
screen "2005_ProNet temperature input" 1280x800, template "Navigation"
   Group "Group" at 118,204 size 1041x515
   TextField "Text field_3" at 172,348 size 56x25; Text 'Mode'
   TextField "Text field_4" at 172,388 size 56x25; Text 'Mode'
   TextField "Text field_5" at 172,430 size 105x25; Text 'Value_10V'
   TextField "Text field_6" at 172,470 size 139x25; Text 'Tank_Average'
   TextField "Text field_7" at 457,550 size 254x25; Text '0:0.. 5 V; 1: -5.. +5 V;'
   TextField "Text field_8" at 702,550 size 308x25; Text '2:0.. 10 V; 3: -10 V.. +10 V;'
   TextField "Text field_9" at 222,550 size 56x25; Text 'Mode'
   TextField "Text field_11" at 222,606 size 105x25; Text 'Value_10V'
   TextField "Text field_12" at 222,634 size 139x25; Text 'Tank_Average'
   TextField "Text field_14" at 457,606 size 366x25; Text 'Max Value for input 10V or 138.5 ohm'
   TextField "Text field_15" at 456,634 size 222x25; Text 'Time for average [ms]'
   TextField "Text field_16" at 373,302 size 46x25; Text '1'
   TextField "Text field_17" at 469,302 size 46x25; Text '2'
   TextField "Text field_18" at 565,302 size 46x25; Text '3'
   TextField "Text field_19" at 661,302 size 46x25; Text '4'
   TextField "Text field_20" at 757,302 size 46x25; Text '5'
   TextField "Text field_21" at 853,302 size 46x25; Text '6'
   TextField "Text field_22" at 949,302 size 46x25; Text '7'
   TextField "Text field_23" at 1045,302 size 46x25; Text '8'
   SymbolicIOField "Symbolic I/O field_5" at 326,104 size 451x32; TextOn '1'; TextOff '0'; TextList "Pronet_Analog_Input"
      ProcessValue <- "PN_AI_SetIndex"
   Button "b_Incress_PronetAnalogInput" at 787,104 size 46x32; TextOff 'Text'; PictureOff "NEXT"
      on Press: function_dd21b452("PN_AI_SetIndex", 1)
   Button "b_Decress_PronetAnalogInput" at 270,104 size 46x32; TextOff 'Text'; PictureOff "BEFORE"
      on Press: function_b9b71300("PN_AI_SetIndex", 1)
   Button "Button_1" at 1017,244 size 96x32; TextOff 'Active'
      on Press: InvertBit("PN_AI_Module{0}_AIResistive_8_Active")
      Appearance <- "PN_AI_Module{0}_AIResistive_8_Active"
   TextField "Text field_1" at 428,145 size 247x29; Text 'ProNet Configuration'
   IOField "Pronet_Analog_Input/Mode1" at 341,344 size 80x32; FormatPattern 9999999
      ProcessValue <- "PN_AI_Module{0}_AI8_X14_0_Data_Data[1]_Betriebsart"
   IOField "I/O field_2" at 437,344 size 80x32; FormatPattern 9999999
      ProcessValue <- "PN_AI_Module{0}_AI8_X14_0_Data_Data[2]_Betriebsart"
   IOField "I/O field_3" at 533,344 size 80x32; FormatPattern 9999999
      ProcessValue <- "PN_AI_Module{0}_AI8_X14_0_Data_Data[3]_Betriebsart"
   IOField "I/O field_4" at 629,344 size 80x32; FormatPattern 9999999
      ProcessValue <- "PN_AI_Module{0}_AI8_X14_0_Data_Data[4]_Betriebsart"
   IOField "I/O field_5" at 725,344 size 80x32; FormatPattern 9999999
      ProcessValue <- "PN_AI_Module{0}_AI8_X14_0_Data_Data[5]_Betriebsart"
   IOField "I/O field_6" at 821,344 size 80x32; FormatPattern 9999999
      ProcessValue <- "PN_AI_Module{0}_AI8_X14_0_Data_Data[6]_Betriebsart"
   IOField "I/O field_7" at 917,344 size 80x32; FormatPattern 9999999
      ProcessValue <- "PN_AI_Module{0}_AI8_X14_0_Data_Data[7]_Betriebsart"
   IOField "I/O field_8" at 1013,344 size 80x32; FormatPattern 9999999
      ProcessValue <- "PN_AI_Module{0}_AI8_X14_0_Data_Data[8]_Betriebsart"
   IOField "I/O field_9" at 341,384 size 80x32; FormatPattern 9999999
      ProcessValue <- "PN_AI_Module{0}_AIResistive_8_TemperatureInput_Data{1}_Einheit"
   IOField "I/O field_10" at 437,384 size 80x32; FormatPattern 9999999
      ProcessValue <- "PN_AI_Module{0}_AIResistive_8_TemperatureInput_Data{2}_Einheit"
   IOField "I/O field_11" at 533,384 size 80x32; FormatPattern 9999999
      ProcessValue <- "PN_AI_Module{0}_AIResistive_8_TemperatureInput_Data{3}_Einheit"
   IOField "I/O field_12" at 629,384 size 80x32; FormatPattern 9999999
      ProcessValue <- "PN_AI_Module{0}_AIResistive_8_TemperatureInput_Data{4}_Einheit"
   IOField "I/O field_13" at 725,384 size 80x32; FormatPattern 9999999
      ProcessValue <- "PN_AI_Module{0}_AIResistive_8_TemperatureInput_Data{5}_Einheit"
   IOField "I/O field_14" at 821,384 size 80x32; FormatPattern 9999999
      ProcessValue <- "PN_AI_Module{0}_AIResistive_8_TemperatureInput_Data{6}_Einheit"
   IOField "I/O field_15" at 917,384 size 80x32; FormatPattern 9999999
      ProcessValue <- "PN_AI_Module{0}_AIResistive_8_TemperatureInput_Data{7}_Einheit"
   IOField "I/O field_16" at 1013,384 size 80x32; FormatPattern 9999999
      ProcessValue <- "PN_AI_Module{0}_AIResistive_8_TemperatureInput_Data{8}_Einheit"
   IOField "I/O field_17" at 341,426 size 80x32; FormatPattern 9999999
      ProcessValue <- "PN_AI_Module{0}_AIResistive_8_TemperatureInput_Data{1}_ErsatzwertDrahtbruch"
   IOField "I/O field_18" at 437,426 size 80x32; FormatPattern 9999999
      ProcessValue <- "PN_AI_Module{0}_AIResistive_8_TemperatureInput_Data{2}_ErsatzwertDrahtbruch"
   IOField "I/O field_19" at 533,426 size 80x32; FormatPattern 9999999
      ProcessValue <- "PN_AI_Module{0}_AIResistive_8_TemperatureInput_Data{3}_ErsatzwertDrahtbruch"
   IOField "I/O field_20" at 629,426 size 80x32; FormatPattern 9999999
      ProcessValue <- "PN_AI_Module{0}_AIResistive_8_TemperatureInput_Data{4}_ErsatzwertDrahtbruch"
   IOField "I/O field_21" at 725,426 size 80x32; FormatPattern 9999999
      ProcessValue <- "PN_AI_Module{0}_AIResistive_8_TemperatureInput_Data{5}_ErsatzwertDrahtbruch"
   IOField "I/O field_22" at 821,426 size 80x32; FormatPattern 9999999
      ProcessValue <- "PN_AI_Module{0}_AIResistive_8_TemperatureInput_Data{6}_ErsatzwertDrahtbruch"
   IOField "I/O field_23" at 917,426 size 80x32; FormatPattern 9999999
      ProcessValue <- "PN_AI_Module{0}_AIResistive_8_TemperatureInput_Data{7}_ErsatzwertDrahtbruch"
   IOField "I/O field_24" at 1013,426 size 80x32; FormatPattern 9999999
      ProcessValue <- "PN_AI_Module{0}_AIResistive_8_TemperatureInput_Data{8}_ErsatzwertDrahtbruch"
   IOField "I/O field_25" at 341,466 size 80x32; FormatPattern 9999999
      ProcessValue <- "PN_AI_Module{0}_AIResistive_8_TemperatureInput_Data{1}_Mittelwertzeit"
   IOField "I/O field_26" at 437,466 size 80x32; FormatPattern 9999999
      ProcessValue <- "PN_AI_Module{0}_AIResistive_8_TemperatureInput_Data{2}_Mittelwertzeit"
   IOField "I/O field_27" at 533,466 size 80x32; FormatPattern 9999999
      ProcessValue <- "PN_AI_Module{0}_AIResistive_8_TemperatureInput_Data{3}_Mittelwertzeit"
   IOField "I/O field_28" at 629,466 size 80x32; FormatPattern 9999999
      ProcessValue <- "PN_AI_Module{0}_AIResistive_8_TemperatureInput_Data{4}_Mittelwertzeit"
   IOField "I/O field_29" at 725,466 size 80x32; FormatPattern 9999999
      ProcessValue <- "PN_AI_Module{0}_AIResistive_8_TemperatureInput_Data{5}_Mittelwertzeit"
   IOField "I/O field_30" at 821,466 size 80x32; FormatPattern 9999999
      ProcessValue <- "PN_AI_Module{0}_AIResistive_8_TemperatureInput_Data{6}_Mittelwertzeit"
   IOField "I/O field_31" at 917,466 size 80x32; FormatPattern 9999999
      ProcessValue <- "PN_AI_Module{0}_AIResistive_8_TemperatureInput_Data{7}_Mittelwertzeit"
   IOField "I/O field_32" at 1013,466 size 80x32; FormatPattern 9999999
      ProcessValue <- "PN_AI_Module{0}_AIResistive_8_TemperatureInput_Data{8}_Mittelwertzeit"
   IOField "I/O field_33" at 1017,159 size 96x32; FormatPattern 99999
      ProcessValue <- "PN_AI_Module{0}_AIResistive_8_Address"
   TextField "Text field_2" at 888,162 size 122x25; Text 'Start Adress'
   TextField "Text field_24" at 460,576 size 71x25; Text '0...100'
   TextField "Text field_25" at 524,576 size 36x18; Text 'o'
   TextField "Text field_26" at 533,576 size 46x25; Text 'C'
   TextField "Text field_27" at 554,576 size 49x25; Text '-100'
   TextField "Text field_28" at 595,576 size 36x18; Text 'o'
   TextField "Text field_29" at 604,576 size 46x25; Text 'C'
   TextField "Text field_30" at 617,576 size 74x25; Text '...+100'
   TextField "Text field_31" at 681,576 size 36x18; Text 'o'
   TextField "Text field_32" at 690,576 size 46x25; Text 'C'
   TextField "Text field_36" at 716,576 size 71x25; Text '0...200'
   TextField "Text field_37" at 776,576 size 36x18; Text 'o'
   TextField "Text field_38" at 785,576 size 46x25; Text 'C'
   TextField "Text field_39" at 814,576 size 49x25; Text '-200'
   TextField "Text field_40" at 855,576 size 36x18; Text 'o'
   TextField "Text field_41" at 864,576 size 46x25; Text 'C'
   TextField "Text field_42" at 877,576 size 74x25; Text '...+200'
   TextField "Text field_43" at 941,576 size 36x18; Text 'o'
   TextField "Text field_44" at 950,576 size 46x25; Text 'C'
   TextField "Text field_10" at 476,270 size 149x29; Text 'Analog input'

screen "2002_ProNet Flow control" 1280x800, template "Navigation"
   on GenerateScreen: SetBit("PN_FlowRate_Component{0}_FlowC_F_Hardware_Request"); SetBit("PN_FlowRate_Component{0}_FlowC_F_GeneralParameters_Request"); SetBit("PN_FlowRate_Component{0}_FlowC_F_Grenzen_Request"); SetBit("PN_FlowRate_Component{0}_FlowC_F_SkalierungAI_Request")
   Group "Group" at 118,168 size 1041x597
   TextField "Text field_2" at 439,140 size 225x27; Text 'Pronet Configuration'
   TextField "Text field_3" at 797,199 size 128x25; Text 'Start Adress'
   TextField "Text field_4" at 168,244 size 100x27; Text 'General :'
   TextField "Text field_5" at 271,273 size 266x25; Text 'Calibration [0,0001 g/Imp]'
   TextField "Text field_6" at 271,307 size 248x25; Text 'Maximum flow [0,01 g/s]'
   TextField "Text field_7" at 271,342 size 276x25; Text 'Close loop control time [Ms]'
   TextField "Text field_8" at 271,376 size 289x25; Text 'time for moving average [ms]'
   TextField "Text field_9" at 168,413 size 129x27; Text 'Delimiting :'
   TextField "Text field_10" at 271,450 size 431x25; Text 'Upper limit manipulated variable (0.0 ... 1.0)'
   TextField "Text field_11" at 271,484 size 440x25; Text 'Lower limit manipulated variable (-1.0 ... 1.0)'
   TextField "Text field_12" at 271,519 size 551x25; Text 'Time delay warning max. voltage limit (0.001 ... 10.0) [s]'
   TextField "Text field_13" at 271,553 size 547x25; Text 'Time delay warning min. voltage limit (0.00q ... 10.0) [s] / Time delay warning min. voltage limit (0.001 ... 10.0) [s]'
   TextField "Text field_14" at 168,590 size 304x27; Text 'Analog input values for FPB:'
   TextField "Text field_15" at 271,623 size 407x25; Text 'Maximum output voltage (100 ... +32767)'
   TextField "Text field_16" at 271,655 size 435x25; Text 'Minimum output voltage (-32767 ... +32767)'
   TextField "Text field_17" at 271,687 size 272x25; Text 'time for moving average [s]'
   SymbolicIOField "Symbolic I/O field_5" at 326,104 size 451x32; TextOn '1'; TextOff '0'; TextList "Pump_Name"
      ProcessValue <- "PN_FlowRate_SetIndex"
   Button "b_Increass_Pronet_FlowControl" at 786,104 size 46x32; TextOff 'Text'; PictureOff "NEXT"
      on Press: function_dd21b452("PN_FlowRate_SetIndex", 1)
   Button "b_Decress_PronetFlowControl" at 272,104 size 46x32; TextOff 'Text'; PictureOff "BEFORE"
      on Press: function_b9b71300("PN_FlowRate_SetIndex", 1)
   IOField "Pronet_FlowControl_AnaIn_Max_InputVoltage" at 776,616 size 96x32; FormatPattern 9999.999
      ProcessValue <- "PN_FlowRate_Component{0}_FlowC_F_SkalierungAI_Data_Bereichsobergrenze"
   IOField "I/O field_2" at 776,651 size 96x32; FormatPattern s9999.999
      ProcessValue <- "PN_FlowRate_Component{0}_FlowC_F_SkalierungAI_Data_Bereichsuntergrenze"
   IOField "I/O field_3" at 776,687 size 96x32; FormatPattern 9999.999
      ProcessValue <- "PN_FlowRate_Component{0}_FlowC_F_SkalierungAI_Data_Mittelwertzeit"
   IOField "I/O field_4" at 935,198 size 96x32; FormatPattern 9999
      ProcessValue <- "PN_FlowRate_Component{0}_FlowC_F_Address"
      on OnFinishInput: SetBit("PN_FlowRate_Component{0}_FlowC_F_Hardware_Request"); SetBit("PN_FlowRate_Component{0}_FlowC_F_GeneralParameters_Request"); SetBit("PN_FlowRate_Component{0}_FlowC_F_Grenzen_Request"); SetBit("PN_FlowRate_Component{0}_FlowC_F_SkalierungAI_Request")
   Button "Button_1" at 1038,198 size 96x32; TextOff 'Active'
      on Press: InvertBit("PN_FlowRate_Component{0}_FlowC_F_Active")
      Appearance <- "PN_FlowRate_Component{0}_FlowC_F_Active"
   IOField "I/O field_5" at 776,372 size 96x32; FormatPattern 9999.999
      ProcessValue <- "PN_FlowRate_Component{0}_FlowC_F_GeneralParameters_Data_Filterzeit"
   IOField "I/O field_6" at 776,446 size 96x32; FormatPattern 9.999
      ProcessValue <- "PN_FlowRate_Component{0}_FlowC_F_Grenzen_Data_ObergrenzeStellgröße"
   IOField "I/O field_7" at 776,480 size 96x32; FormatPattern 9.999
      ProcessValue <- "PN_FlowRate_Component{0}_FlowC_F_Grenzen_Data_UntergrenzeStellgröße"
   IOField "I/O field_8" at 776,515 size 96x32; FormatPattern 99.999
      ProcessValue <- "PN_FlowRate_Component{0}_FlowC_F_Grenzen_Data_VerzögerungAlarmObergrenze"
   IOField "I/O field_9" at 776,549 size 96x32; FormatPattern 99.999
      ProcessValue <- "PN_FlowRate_Component{0}_FlowC_F_Grenzen_Data_VerzögerungAlarmUntergrenze"
   IOField "I/O field_10" at 776,269 size 96x32; FormatPattern s9999.999
      ProcessValue <- "PN_FlowRate_Component{0}_FlowC_F_GeneralParameters_Data_Kalibrierfaktor"
   IOField "I/O field_11" at 776,303 size 96x32; FormatPattern s9999.99
      ProcessValue <- "PN_FlowRate_Component{0}_FlowC_F_GeneralParameters_Data_MaxDurchfluss"
   IOField "I/O field_12" at 776,338 size 96x32; FormatPattern 9999.999
      ProcessValue <- "PN_FlowRate_Component{0}_FlowC_F_GeneralParameters_Data_Nachstellzeit"
   TextField "Text field_1" at 483,198 size 137x27; Text 'Flow control'

screen "2006_ProNet Nozzle configuration" 1280x800, template "Navigation"
   on GenerateScreen: SetBit("PN_Mixinghead_Send"); SetBit("PN_Mixinghead_Mixinghead{0}_Digital_GeneralParameters_Request")
   Group "Group" at 100,196 size 1078x475
   TextField "Text field_4" at 105,334 size 46x25; Text 'Text'
   TextField "Text field_9" at 364,282 size 101x20; Text 'Start Adress'
   TextField "Text field_10" at 472,274 size 145x36; Text 'Mixinghead change Mixinghead channel'
   TextField "Text field_11" at 608,274 size 156x36; Text 'Mixhead vlve output Output for nozzle'
   TextField "Text field_12" at 746,274 size 127x36; Text 'Proximity switch Polarity of nozzle'
   TextField "Text field_13" at 886,274 size 126x36; Text 'External release Output for bypass'
   TextField "Text field_14" at 1025,274 size 127x36; Text 'Proximity switch Polarity of bypass'
   Button "Button_1" at 264,329 size 88x27; TextOff 'Active'
      on Press: InvertBit("PN_Mixinghead_Mixinghead{0}_DüseBypass{1}_Active")
      Appearance <- "PN_Mixinghead_Mixinghead{0}_DüseBypass{1}_Active"
   TextField "Text field_1" at 428,142 size 247x29; Text 'ProNet Configuration'
   SymbolicIOField "Symbolic I/O field_5" at 326,104 size 451x32; TextOn '1'; TextOff '0'; TextList "MH_NO"
      ProcessValue <- "PN_Mixinghead_SetIndex"
   Button "Pronet_Increass_Nozzle1" at 786,104 size 46x32; TextOff 'Text'; PictureOff "NEXT"
      on Press: function_dd21b452("PN_Mixinghead_SetIndex", 1); SetBit("PN_Mixinghead_Send")
   Button "Pronet_Decress_Nozzle1" at 271,104 size 46x32; TextOff 'Text'; PictureOff "BEFORE"
      on Press: function_b9b71300("PN_Mixinghead_SetIndex", 1); SetBit("PN_Mixinghead_Send")
   IOField "Pronet_Nozzle1_StartAdress" at 366,327 size 96x32; FormatPattern 99999
      ProcessValue <- "PN_Mixinghead_Mixinghead{0}_DüseBypass{1}_Address"
   IOField "I/O field_2" at 366,374 size 96x32; FormatPattern 99999
      ProcessValue <- "PN_Mixinghead_Mixinghead{0}_DüseBypass{2}_Address"
   IOField "I/O field_3" at 366,420 size 96x32; FormatPattern 99999
      ProcessValue <- "PN_Mixinghead_Mixinghead{0}_DüseBypass{3}_Address"
   IOField "I/O field_4" at 366,465 size 96x32; FormatPattern 99999
      ProcessValue <- "PN_Mixinghead_Mixinghead{0}_DüseBypass{4}_Address"
   IOField "I/O field_5" at 366,510 size 96x32; FormatPattern 99999
      ProcessValue <- "PN_Mixinghead_Mixinghead{0}_DüseBypass{5}_Address"
   IOField "I/O field_6" at 366,554 size 96x32; FormatPattern 99999
      ProcessValue <- "PN_Mixinghead_Mixinghead{0}_DüseBypass{6}_Address"
   SymbolicIOField "Symbolic I/O field_1" at 472,327 size 128x32; TextOff '0'; TextOn '1'; TextList "Pronet_Mixinghead Chanel"
      ProcessValue <- "PN_Mixinghead_Mixinghead{0}_DüseBypass{1}_Visualisierung_MHChannel"
   SymbolicIOField "Symbolic I/O field_2" at 472,374 size 128x32; TextOn '1'; TextOff '0'; TextList "Pronet_Mixinghead Chanel"
      ProcessValue <- "PN_Mixinghead_Mixinghead{0}_DüseBypass{2}_Visualisierung_MHChannel"
   SymbolicIOField "Symbolic I/O field_3" at 472,420 size 128x32; TextOn '1'; TextOff '0'; TextList "Pronet_Mixinghead Chanel"
      ProcessValue <- "PN_Mixinghead_Mixinghead{0}_DüseBypass{3}_Visualisierung_MHChannel"
   SymbolicIOField "Symbolic I/O field_4" at 472,465 size 128x32; TextOn '1'; TextOff '0'; TextList "Pronet_Mixinghead Chanel"
      ProcessValue <- "PN_Mixinghead_Mixinghead{0}_DüseBypass{4}_Visualisierung_MHChannel"
   SymbolicIOField "Symbolic I/O field_6" at 472,510 size 128x32; TextOn '1'; TextOff '0'; TextList "Pronet_Mixinghead Chanel"
      ProcessValue <- "PN_Mixinghead_Mixinghead{0}_DüseBypass{5}_Visualisierung_MHChannel"
   SymbolicIOField "Symbolic I/O field_7" at 472,554 size 128x32; TextOn '1'; TextOff '0'; TextList "Pronet_Mixinghead Chanel"
      ProcessValue <- "PN_Mixinghead_Mixinghead{0}_DüseBypass{6}_Visualisierung_MHChannel"
   SymbolicIOField "Symbolic I/O field_8" at 608,327 size 128x32; TextOn '1'; TextOff '0'; TextList "Pronet_Mixinghead_Output_Valve_Numb"
      ProcessValue <- "PN_Mixinghead_Mixinghead{0}_DüseBypass{1}_Visualisierung_OutputForNozzle"
   SymbolicIOField "Symbolic I/O field_9" at 608,374 size 128x32; TextOn '1'; TextOff '0'; TextList "Pronet_Mixinghead_Output_Valve_Numb"
      ProcessValue <- "PN_Mixinghead_Mixinghead{0}_DüseBypass{2}_Visualisierung_OutputForNozzle"
   SymbolicIOField "Symbolic I/O field_10" at 608,420 size 128x32; TextOn '1'; TextOff '0'; TextList "Pronet_Mixinghead_Output_Valve_Numb"
      ProcessValue <- "PN_Mixinghead_Mixinghead{0}_DüseBypass{3}_Visualisierung_OutputForNozzle"
   SymbolicIOField "Symbolic I/O field_11" at 608,465 size 128x32; TextOn '1'; TextOff '0'; TextList "Pronet_Mixinghead_Output_Valve_Numb"
      ProcessValue <- "PN_Mixinghead_Mixinghead{0}_DüseBypass{4}_Visualisierung_OutputForNozzle"
   SymbolicIOField "Symbolic I/O field_12" at 608,510 size 128x32; TextOn '1'; TextOff '0'; TextList "Pronet_Mixinghead_Output_Valve_Numb"
      ProcessValue <- "PN_Mixinghead_Mixinghead{0}_DüseBypass{5}_Visualisierung_OutputForNozzle"
   SymbolicIOField "Symbolic I/O field_13" at 608,554 size 128x32; TextOn '1'; TextOff '0'; TextList "Pronet_Mixinghead_Output_Valve_Numb"
      ProcessValue <- "PN_Mixinghead_Mixinghead{0}_DüseBypass{6}_Visualisierung_OutputForNozzle"
   SymbolicIOField "Symbolic I/O field_14" at 886,327 size 128x32; TextOn '1'; TextOff '0'; TextList "Pronet_Mixinghead_Output_Valve_Numb"
      ProcessValue <- "PN_Mixinghead_Mixinghead{0}_DüseBypass{1}_Visualisierung_OutputForBypass"
   SymbolicIOField "Symbolic I/O field_15" at 886,374 size 128x32; TextOn '1'; TextOff '0'; TextList "Pronet_Mixinghead_Output_Valve_Numb"
      ProcessValue <- "PN_Mixinghead_Mixinghead{0}_DüseBypass{2}_Visualisierung_OutputForBypass"
   SymbolicIOField "Symbolic I/O field_16" at 886,420 size 128x32; TextOn '1'; TextOff '0'; TextList "Pronet_Mixinghead_Output_Valve_Numb"
      ProcessValue <- "PN_Mixinghead_Mixinghead{0}_DüseBypass{3}_Visualisierung_OutputForBypass"
   SymbolicIOField "Symbolic I/O field_17" at 886,465 size 128x32; TextOn '1'; TextOff '0'; TextList "Pronet_Mixinghead_Output_Valve_Numb"
      ProcessValue <- "PN_Mixinghead_Mixinghead{0}_DüseBypass{4}_Visualisierung_OutputForBypass"
   SymbolicIOField "Symbolic I/O field_18" at 886,510 size 128x32; TextOn '1'; TextOff '0'; TextList "Pronet_Mixinghead_Output_Valve_Numb"
      ProcessValue <- "PN_Mixinghead_Mixinghead{0}_DüseBypass{5}_Visualisierung_OutputForBypass"
   SymbolicIOField "Symbolic I/O field_19" at 886,554 size 128x32; TextOn '1'; TextOff '0'; TextList "Pronet_Mixinghead_Output_Valve_Numb"
      ProcessValue <- "PN_Mixinghead_Mixinghead{0}_DüseBypass{6}_Visualisierung_OutputForBypass"
   SymbolicIOField "Symbolic I/O field_20" at 746,327 size 128x32; TextOn '1'; TextOff '0'; TextList "Pronet_NO_NC"
      ProcessValue <- "PN_Mixinghead_Mixinghead{0}_DüseBypass{1}_Visualisierung_PolarityNozzle"
   SymbolicIOField "Symbolic I/O field_21" at 746,374 size 128x32; TextOn '1'; TextOff '0'; TextList "Pronet_NO_NC"
      ProcessValue <- "PN_Mixinghead_Mixinghead{0}_DüseBypass{2}_Visualisierung_PolarityNozzle"
   SymbolicIOField "Symbolic I/O field_22" at 746,420 size 128x32; TextOn '1'; TextOff '0'; TextList "Pronet_NO_NC"
      ProcessValue <- "PN_Mixinghead_Mixinghead{0}_DüseBypass{3}_Visualisierung_PolarityNozzle"
   SymbolicIOField "Symbolic I/O field_23" at 746,465 size 128x32; TextOn '1'; TextOff '0'; TextList "Pronet_NO_NC"
      ProcessValue <- "PN_Mixinghead_Mixinghead{0}_DüseBypass{4}_Visualisierung_PolarityNozzle"
   SymbolicIOField "Symbolic I/O field_24" at 746,510 size 128x32; TextOn '1'; TextOff '0'; TextList "Pronet_NO_NC"
      ProcessValue <- "PN_Mixinghead_Mixinghead{0}_DüseBypass{5}_Visualisierung_PolarityNozzle"
   SymbolicIOField "Symbolic I/O field_25" at 746,554 size 128x32; TextOn '1'; TextOff '0'; TextList "Pronet_NO_NC"
      ProcessValue <- "PN_Mixinghead_Mixinghead{0}_DüseBypass{6}_Visualisierung_PolarityNozzle"
   SymbolicIOField "Symbolic I/O field_26" at 1025,327 size 128x32; TextOn '1'; TextOff '0'; TextList "Pronet_NO_NC"
      ProcessValue <- "PN_Mixinghead_Mixinghead{0}_DüseBypass{1}_Visualisierung_PolarityBypass"
   SymbolicIOField "Symbolic I/O field_27" at 1025,374 size 128x32; TextOn '1'; TextOff '0'; TextList "Pronet_NO_NC"
      ProcessValue <- "PN_Mixinghead_Mixinghead{0}_DüseBypass{2}_Visualisierung_PolarityBypass"
   SymbolicIOField "Symbolic I/O field_28" at 1025,420 size 128x32; TextOn '1'; TextOff '0'; TextList "Pronet_NO_NC"
      ProcessValue <- "PN_Mixinghead_Mixinghead{0}_DüseBypass{3}_Visualisierung_PolarityBypass"
   SymbolicIOField "Symbolic I/O field_29" at 1025,465 size 128x32; TextOn '1'; TextOff '0'; TextList "Pronet_NO_NC"
      ProcessValue <- "PN_Mixinghead_Mixinghead{0}_DüseBypass{4}_Visualisierung_PolarityBypass"
   SymbolicIOField "Symbolic I/O field_30" at 1025,510 size 128x32; TextOn '1'; TextOff '0'; TextList "Pronet_NO_NC"
      ProcessValue <- "PN_Mixinghead_Mixinghead{0}_DüseBypass{5}_Visualisierung_PolarityBypass"
   SymbolicIOField "Symbolic I/O field_31" at 1025,554 size 128x32; TextOn '1'; TextOff '0'; TextList "Pronet_NO_NC"
      ProcessValue <- "PN_Mixinghead_Mixinghead{0}_DüseBypass{6}_Visualisierung_PolarityBypass"
   Button "Button_2" at 264,376 size 88x27; TextOff 'Active'
      on Press: InvertBit("PN_Mixinghead_Mixinghead{0}_DüseBypass{2}_Active")
      Appearance <- "PN_Mixinghead_Mixinghead{0}_DüseBypass{2}_Active"
   Button "Button_3" at 264,422 size 88x27; TextOff 'Active'
      on Press: InvertBit("PN_Mixinghead_Mixinghead{0}_DüseBypass{3}_Active")
      Appearance <- "PN_Mixinghead_Mixinghead{0}_DüseBypass{3}_Active"
   Button "Button_4" at 264,467 size 88x27; TextOff 'Active'
      on Press: InvertBit("PN_Mixinghead_Mixinghead{0}_DüseBypass{4}_Active")
      Appearance <- "PN_Mixinghead_Mixinghead{0}_DüseBypass{4}_Active"
   Button "Button_5" at 264,512 size 88x27; TextOff 'Active'
      on Press: InvertBit("PN_Mixinghead_Mixinghead{0}_DüseBypass{5}_Active")
      Appearance <- "PN_Mixinghead_Mixinghead{0}_DüseBypass{5}_Active"
   Button "Button_6" at 264,556 size 88x27; TextOff 'Active'
      on Press: InvertBit("PN_Mixinghead_Mixinghead{0}_DüseBypass{6}_Active")
      Appearance <- "PN_Mixinghead_Mixinghead{0}_DüseBypass{6}_Active"
   TextField "Text field_2" at 468,219 size 226x29; Text 'Nozzle control / Nozzle cofiguration'
   TextField "Text field_3" at 129,332 size 130x22; Text 'Text'
   TextField "Text field_5" at 129,379 size 130x22; Text 'Text'
   TextField "Text field_6" at 129,425 size 130x22; Text 'Text'
   TextField "Text field_7" at 129,470 size 130x22; Text 'Text'
   TextField "Text field_8" at 129,515 size 130x22; Text 'Text'
   TextField "Text field_15" at 129,559 size 130x22; Text 'Text'

screen "2007_ProNet Nozzle times" 1280x800, template "Navigation"
   on GenerateScreen: SetBit("PN_Mixinghead_Send"); SetBit("PN_Mixinghead_Mixinghead{0}_Digital_GeneralParameters_Request")
   Group "Group" at 118,195 size 1041x469
   TextField "Text field_1" at 428,143 size 247x29; Text 'ProNet Configuration'
   SymbolicIOField "Symbolic I/O field_5" at 326,104 size 451x32; TextOn '1'; TextOff '0'; TextList "MH_NO"
      ProcessValue <- "PN_Mixinghead_SetIndex"
   Button "b_Incress_Pronet_NozzleControl" at 787,104 size 46x32; TextOff 'Text'; PictureOff "NEXT"
      on Press: function_dd21b452("PN_Mixinghead_SetIndex", 1); SetBit("PN_Mixinghead_Send")
   Button "b_Decress_Pronet_NozzleControl" at 269,104 size 46x32; TextOff 'Text'; PictureOff "BEFORE"
      on Press: function_b9b71300("PN_Mixinghead_SetIndex", 1); SetBit("PN_Mixinghead_Send")
   TextField "Text field_3" at 151,332 size 213x22; Text 'Text'
   TextField "Text field_5" at 151,379 size 213x22; Text 'Text'
   TextField "Text field_6" at 151,425 size 213x22; Text 'Text'
   TextField "Text field_7" at 151,470 size 213x22; Text 'Text'
   TextField "Text field_8" at 151,515 size 213x22; Text 'Text'
   TextField "Text field_15" at 151,559 size 213x22; Text 'Text'
   TextField "Text field_2" at 506,332 size 42x22; Text '[s]'
   IOField "Time1_NozzleControl" at 402,327 size 96x32; FormatPattern 9999.999
      ProcessValue <- "PN_Mixinghead_Mixinghead{0}_DüseBypass{1}_Zeiten_Data_ÜberlappungD_B"
   IOField "I/O field_2" at 584,327 size 96x32; FormatPattern 9999.999
      ProcessValue <- "PN_Mixinghead_Mixinghead{0}_DüseBypass{1}_Zeiten_Data_ÜberlappungB_D"
   IOField "I/O field_3" at 763,327 size 96x32; FormatPattern 9999.999
      ProcessValue <- "PN_Mixinghead_Mixinghead{0}_DüseBypass{1}_Zeiten_Data_VerzögerungSchussstart"
   IOField "I/O field_4" at 945,327 size 96x32; FormatPattern 9999.999
      ProcessValue <- "PN_Mixinghead_Mixinghead{0}_DüseBypass{1}_Zeiten_Data_VerzögerungSchussende"
   IOField "I/O field_5" at 402,374 size 96x32; FormatPattern 9999.999
      ProcessValue <- "PN_Mixinghead_Mixinghead{0}_DüseBypass{2}_Zeiten_Data_ÜberlappungD_B"
   IOField "I/O field_6" at 584,374 size 96x32; FormatPattern 9999.999
      ProcessValue <- "PN_Mixinghead_Mixinghead{0}_DüseBypass{2}_Zeiten_Data_ÜberlappungB_D"
   IOField "I/O field_7" at 763,374 size 96x32; FormatPattern 9999.999
      ProcessValue <- "PN_Mixinghead_Mixinghead{0}_DüseBypass{2}_Zeiten_Data_VerzögerungSchussstart"
   IOField "I/O field_8" at 945,374 size 96x32; FormatPattern 9999.999
      ProcessValue <- "PN_Mixinghead_Mixinghead{0}_DüseBypass{2}_Zeiten_Data_VerzögerungSchussende"
   IOField "I/O field_9" at 402,420 size 96x32; FormatPattern 9999.999
      ProcessValue <- "PN_Mixinghead_Mixinghead{0}_DüseBypass{3}_Zeiten_Data_ÜberlappungD_B"
   IOField "I/O field_10" at 584,420 size 96x32; FormatPattern 9999.999
      ProcessValue <- "PN_Mixinghead_Mixinghead{0}_DüseBypass{3}_Zeiten_Data_ÜberlappungB_D"
   IOField "I/O field_11" at 763,420 size 96x32; FormatPattern 9999.999
      ProcessValue <- "PN_Mixinghead_Mixinghead{0}_DüseBypass{3}_Zeiten_Data_VerzögerungSchussstart"
   IOField "I/O field_12" at 945,420 size 96x32; FormatPattern 9999.999
      ProcessValue <- "PN_Mixinghead_Mixinghead{0}_DüseBypass{3}_Zeiten_Data_VerzögerungSchussende"
   IOField "I/O field_13" at 402,465 size 96x32; FormatPattern 9999.999
      ProcessValue <- "PN_Mixinghead_Mixinghead{0}_DüseBypass{4}_Zeiten_Data_ÜberlappungD_B"
   IOField "I/O field_14" at 584,465 size 96x32; FormatPattern 9999.999
      ProcessValue <- "PN_Mixinghead_Mixinghead{0}_DüseBypass{4}_Zeiten_Data_ÜberlappungB_D"
   IOField "I/O field_15" at 763,465 size 96x32; FormatPattern 9999.999
      ProcessValue <- "PN_Mixinghead_Mixinghead{0}_DüseBypass{4}_Zeiten_Data_VerzögerungSchussstart"
   IOField "I/O field_16" at 945,465 size 96x32; FormatPattern 9999.999
      ProcessValue <- "PN_Mixinghead_Mixinghead{0}_DüseBypass{4}_Zeiten_Data_VerzögerungSchussende"
   IOField "I/O field_17" at 402,510 size 96x32; FormatPattern 9999.999
      ProcessValue <- "PN_Mixinghead_Mixinghead{0}_DüseBypass{5}_Zeiten_Data_ÜberlappungD_B"
   IOField "I/O field_18" at 584,510 size 96x32; FormatPattern 9999.999
      ProcessValue <- "PN_Mixinghead_Mixinghead{0}_DüseBypass{5}_Zeiten_Data_ÜberlappungB_D"
   IOField "I/O field_19" at 763,510 size 96x32; FormatPattern 9999.999
      ProcessValue <- "PN_Mixinghead_Mixinghead{0}_DüseBypass{5}_Zeiten_Data_VerzögerungSchussstart"
   IOField "I/O field_20" at 945,510 size 96x32; FormatPattern 9999.999
      ProcessValue <- "PN_Mixinghead_Mixinghead{0}_DüseBypass{5}_Zeiten_Data_VerzögerungSchussende"
   IOField "I/O field_21" at 402,554 size 96x32; FormatPattern 9999.999
      ProcessValue <- "PN_Mixinghead_Mixinghead{0}_DüseBypass{6}_Zeiten_Data_ÜberlappungD_B"
   IOField "Pronet_Time2_last" at 584,554 size 96x32; FormatPattern 9999.999
      ProcessValue <- "PN_Mixinghead_Mixinghead{0}_DüseBypass{6}_Zeiten_Data_ÜberlappungB_D"
   IOField "I/O field_23" at 763,554 size 96x32; FormatPattern 9999.999
      ProcessValue <- "PN_Mixinghead_Mixinghead{0}_DüseBypass{6}_Zeiten_Data_VerzögerungSchussstart"
   IOField "I/O field_24" at 945,554 size 96x32; FormatPattern 9999.999
      ProcessValue <- "PN_Mixinghead_Mixinghead{0}_DüseBypass{6}_Zeiten_Data_VerzögerungSchussende"
   TextField "Text field_4" at 417,278 size 115x40; Text 'Time 1 Overlap time D -> B'
   TextField "Text field_9" at 599,278 size 115x40; Text 'Time 2 Overlap time B -> D'
   TextField "Text field_10" at 778,278 size 96x40; Text 'Time 3 Delay time Opening'
   TextField "Text field_11" at 960,278 size 96x40; Text 'Time 4 Delay time Closing'
   TextField "Text field_12" at 506,379 size 42x22; Text '[s]'
   TextField "Text field_13" at 506,425 size 42x22; Text '[s]'
   TextField "Text field_14" at 506,470 size 42x22; Text '[s]'
   TextField "Text field_16" at 506,515 size 42x22; Text '[s]'
   TextField "Text field_17" at 506,559 size 42x22; Text '[s]'
   TextField "Text field_18" at 688,332 size 42x22; Text '[s]'
   TextField "Text field_19" at 688,379 size 42x22; Text '[s]'
   TextField "Text field_20" at 688,425 size 42x22; Text '[s]'
   TextField "Text field_21" at 688,470 size 42x22; Text '[s]'
   TextField "Text field_22" at 688,515 size 42x22; Text '[s]'
   TextField "Text field_23" at 688,559 size 42x22; Text '[s]'
   TextField "Text field_24" at 867,332 size 42x22; Text '[s]'
   TextField "Text field_25" at 867,383 size 42x22; Text '[s]'
   TextField "Text field_26" at 867,425 size 42x22; Text '[s]'
   TextField "Text field_27" at 867,470 size 42x22; Text '[s]'
   TextField "Text field_28" at 867,515 size 42x22; Text '[s]'
   TextField "Text field_29" at 867,559 size 42x22; Text '[s]'
   TextField "Text field_30" at 1046,332 size 42x22; Text '[s]'
   TextField "Text field_31" at 1046,379 size 42x22; Text '[s]'
   TextField "Text field_32" at 1046,425 size 42x22; Text '[s]'
   TextField "Text field_33" at 1046,470 size 42x22; Text '[s]'
   TextField "Text field_34" at 1046,515 size 42x22; Text '[s]'
   TextField "Text field_35" at 1046,559 size 42x22; Text '[s]'
   TextField "Text field_36" at 468,221 size 238x29; Text 'Nozzle control / Nozzle control times'

screen "2009_ProNet Diagnose IO" 1280x800, template "Navigation"
   Button "Button_3" at 326,104 size 451x32; TextOff '_ProNet Module'
   Circle "Circle_1" at 156,230 size 30x30
      Appearance <- "PN_Error_Module{0}_DO_1"
   Circle "Circle_2" at 184,230 size 30x30
      Appearance <- "PN_Error_Module{0}_DO_1"
   Circle "Circle_3" at 212,230 size 30x30
      Appearance <- "PN_Error_Module{0}_DO_1"
   Circle "Circle_4" at 241,230 size 30x30
      Appearance <- "PN_Error_Module{0}_DO_1"
   Circle "Circle_5" at 269,230 size 30x30
      Appearance <- "PN_Error_Module{0}_DO_1"
   Circle "Circle_6" at 297,230 size 30x30
      Appearance <- "PN_Error_Module{0}_DO_1"
   Circle "Circle_7" at 325,230 size 30x30
      Appearance <- "PN_Error_Module{0}_DO_1"
   Circle "Circle_8" at 353,230 size 30x30
      Appearance <- "PN_Error_Module{0}_DO_1"
   Circle "Circle_9" at 400,230 size 30x30
      Appearance <- "PN_Error_Module{0}_DO_1"
   Circle "Circle_10" at 428,230 size 30x30
      Appearance <- "PN_Error_Module{0}_DO_1"
   Circle "Circle_11" at 456,230 size 30x30
      Appearance <- "PN_Error_Module{0}_DO_1"
   Circle "Circle_12" at 485,230 size 30x30
      Appearance <- "PN_Error_Module{0}_DO_1"
   Circle "Circle_13" at 513,230 size 30x30
      Appearance <- "PN_Error_Module{0}_DO_1"
   Circle "Circle_14" at 541,230 size 30x30
      Appearance <- "PN_Error_Module{0}_DO_1"
   Circle "Circle_15" at 569,230 size 30x30
      Appearance <- "PN_Error_Module{0}_DO_1"
   Circle "Circle_16" at 597,230 size 30x30
      Appearance <- "PN_Error_Module{0}_DO_1"
   Circle "Circle_17" at 644,230 size 30x30
      Appearance <- "PN_Error_Module{0}_DO_1"
   Circle "Circle_18" at 672,230 size 30x30
      Appearance <- "PN_Error_Module{0}_DO_1"
   Circle "Circle_19" at 700,230 size 30x30
      Appearance <- "PN_Error_Module{0}_DO_1"
   Circle "Circle_20" at 729,230 size 30x30
      Appearance <- "PN_Error_Module{0}_DO_1"
   Circle "Circle_21" at 757,230 size 30x30
      Appearance <- "PN_Error_Module{0}_DO_1"
   Circle "Circle_22" at 785,230 size 30x30
      Appearance <- "PN_Error_Module{0}_DO_1"
   Circle "Circle_23" at 813,230 size 30x30
      Appearance <- "PN_Error_Module{0}_DO_1"
   Circle "Circle_24" at 841,230 size 30x30
      Appearance <- "PN_Error_Module{0}_DO_1"
   Circle "Circle_25" at 888,230 size 30x30
      Appearance <- "PN_Error_Module{0}_DO_1"
   Circle "Circle_26" at 916,230 size 30x30
      Appearance <- "PN_Error_Module{0}_DO_1"
   Circle "Circle_27" at 944,230 size 30x30
      Appearance <- "PN_Error_Module{0}_DO_1"
   Circle "Circle_28" at 973,230 size 30x30
      Appearance <- "PN_Error_Module{0}_DO_1"
   Circle "Circle_29" at 1001,230 size 30x30
      Appearance <- "PN_Error_Module{0}_DO_1"
   Circle "Circle_30" at 1029,230 size 30x30
      Appearance <- "PN_Error_Module{0}_DO_1"
   Circle "Circle_31" at 1057,230 size 30x30
      Appearance <- "PN_Error_Module{0}_DO_1"
   Circle "Circle_32" at 1085,230 size 30x30
      Appearance <- "PN_Error_Module{0}_DO_1"
   Circle "Circle_33" at 156,638 size 30x30
      Appearance <- "PN_Error_Module{0}_DO"
   Circle "Circle_34" at 184,638 size 30x30
      Appearance <- "PN_Error_Module{0}_DO"
   Circle "Circle_35" at 212,638 size 30x30
      Appearance <- "PN_Error_Module{0}_DO"
   Circle "Circle_36" at 241,638 size 30x30
      Appearance <- "PN_Error_Module{0}_DO"
   Circle "Circle_37" at 269,638 size 30x30
      Appearance <- "PN_Error_Module{0}_DO"
   Circle "Circle_38" at 297,638 size 30x30
      Appearance <- "PN_Error_Module{0}_DO"
   Circle "Circle_39" at 325,638 size 30x30
      Appearance <- "PN_Error_Module{0}_DO"
   Circle "Circle_40" at 353,638 size 30x30
      Appearance <- "PN_Error_Module{0}_DO"
   Circle "Circle_41" at 400,638 size 30x30
      Appearance <- "PN_Error_Module{0}_DO"
   Circle "Circle_42" at 428,638 size 30x30
      Appearance <- "PN_Error_Module{0}_DO"
   Circle "Circle_43" at 456,638 size 30x30
      Appearance <- "PN_Error_Module{0}_DO"
   Circle "Circle_44" at 485,638 size 30x30
      Appearance <- "PN_Error_Module{0}_DO"
   Circle "Circle_45" at 513,638 size 30x30
      Appearance <- "PN_Error_Module{0}_DO"
   Circle "Circle_46" at 541,638 size 30x30
      Appearance <- "PN_Error_Module{0}_DO"
   Circle "Circle_47" at 569,638 size 30x30
      Appearance <- "PN_Error_Module{0}_DO"
   Circle "Circle_48" at 597,638 size 30x30
      Appearance <- "PN_Error_Module{0}_DO"
   Circle "Circle_49" at 644,638 size 30x30
      Appearance <- "PN_Error_Module{0}_DO"
   Circle "Circle_50" at 672,638 size 30x30
      Appearance <- "PN_Error_Module{0}_DO"
   Circle "Circle_51" at 700,638 size 30x30
      Appearance <- "PN_Error_Module{0}_DO"
   Circle "Circle_52" at 729,638 size 30x30
      Appearance <- "PN_Error_Module{0}_DO"
   Circle "Circle_53" at 757,638 size 30x30
      Appearance <- "PN_Error_Module{0}_DO"
   Circle "Circle_54" at 785,638 size 30x30
      Appearance <- "PN_Error_Module{0}_DO"
   Circle "Circle_55" at 813,638 size 30x30
      Appearance <- "PN_Error_Module{0}_DO"
   Circle "Circle_56" at 841,638 size 30x30
      Appearance <- "PN_Error_Module{0}_DO"
   Circle "Circle_57" at 888,638 size 30x30
      Appearance <- "PN_Error_Module{0}_DO"
   Circle "Circle_58" at 916,638 size 30x30
      Appearance <- "PN_Error_Module{0}_DO"
   Circle "Circle_59" at 944,638 size 30x30
      Appearance <- "PN_Error_Module{0}_DO"
   Circle "Circle_60" at 973,638 size 30x30
      Appearance <- "PN_Error_Module{0}_DO"
   Circle "Circle_61" at 1001,638 size 30x30
      Appearance <- "PN_Error_Module{0}_DO"
   Circle "Circle_62" at 1029,638 size 30x30
      Appearance <- "PN_Error_Module{0}_DO"
   Circle "Circle_63" at 1057,638 size 30x30
      Appearance <- "PN_Error_Module{0}_DO"
   Circle "Circle_64" at 1085,638 size 30x30
      Appearance <- "PN_Error_Module{0}_DO"
   TextField "Text field_1" at 513,325 size 43x22; Text 'AIr1'
   TextField "Text field_2" at 513,352 size 43x22; Text 'AIr2'
   TextField "Text field_3" at 513,379 size 43x22; Text 'AIr3'
   TextField "Text field_4" at 513,406 size 43x22; Text 'AIr4'
   TextField "Text field_5" at 513,463 size 43x22; Text 'AIr5'
   TextField "Text field_6" at 513,490 size 43x22; Text 'AIr6'
   TextField "Text field_7" at 513,517 size 43x22; Text 'AIr7'
   TextField "Text field_8" at 513,544 size 43x22; Text 'AIr8'
   IOField "I/O field_1" at 578,320 size 96x32; FormatPattern s99999
      ProcessValue <- "PN_Error_Module{0}_AIr{1}"
   IOField "I/O field_2" at 578,347 size 96x32; FormatPattern s99999
      ProcessValue <- "PN_Error_Module{0}_AIr{2}"
   IOField "I/O field_3" at 578,374 size 96x32; FormatPattern s99999
      ProcessValue <- "PN_Error_Module{0}_AIr{3}"
   IOField "I/O field_4" at 578,401 size 96x32; FormatPattern s99999
      ProcessValue <- "PN_Error_Module{0}_AIr{4}"
   IOField "I/O field_5" at 578,458 size 96x32; FormatPattern s99999
      ProcessValue <- "PN_Error_Module{0}_AIr{5}"
   IOField "I/O field_6" at 578,485 size 96x32; FormatPattern s99999
      ProcessValue <- "PN_Error_Module{0}_AIr{6}"
   IOField "I/O field_7" at 578,512 size 96x32; FormatPattern s99999
      ProcessValue <- "PN_Error_Module{0}_AIr{7}"
   IOField "I/O field_8" at 578,539 size 96x32; FormatPattern s99999
      ProcessValue <- "PN_Error_Module{0}_AIr{8}"
   TextField "Text field_9" at 261,325 size 42x22; Text 'AI1'
   TextField "Text field_10" at 261,352 size 42x22; Text 'AI2'
   TextField "Text field_11" at 261,379 size 42x22; Text 'AI3'
   TextField "Text field_12" at 261,406 size 42x22; Text 'AI4'
   TextField "Text field_13" at 261,463 size 42x22; Text 'AI5'
   TextField "Text field_14" at 261,490 size 42x22; Text 'AI6'
   TextField "Text field_15" at 261,517 size 42x22; Text 'AI7'
   TextField "Text field_16" at 261,544 size 42x22; Text 'AI8'
   IOField "I/O field_9" at 326,320 size 96x32; FormatPattern s99999
      ProcessValue <- "PN_Error_Module{0}_AI{1}"
   IOField "I/O field_10" at 326,347 size 96x32; FormatPattern s99999
      ProcessValue <- "PN_Error_Module{0}_AI{2}"
   IOField "I/O field_11" at 326,374 size 96x32; FormatPattern s99999
      ProcessValue <- "PN_Error_Module{0}_AI{3}"
   IOField "I/O field_12" at 326,401 size 96x32; FormatPattern s99999
      ProcessValue <- "PN_Error_Module{0}_AI{4}"
   IOField "I/O field_13" at 326,458 size 96x32; FormatPattern s99999
      ProcessValue <- "PN_Error_Module{0}_AI{5}"
   IOField "I/O field_14" at 326,485 size 96x32; FormatPattern s99999
      ProcessValue <- "PN_Error_Module{0}_AI{6}"
   IOField "I/O field_15" at 326,512 size 96x32; FormatPattern s99999
      ProcessValue <- "PN_Error_Module{0}_AI{7}"
   IOField "I/O field_16" at 326,539 size 96x32; FormatPattern s99999
      ProcessValue <- "PN_Error_Module{0}_AI{8}"
   TextField "Text field_17" at 160,258 size 22x53; Text 'DI0.0'
   TextField "Text field_18" at 188,258 size 22x53; Text 'DI0.1'
   TextField "Text field_19" at 216,258 size 22x53; Text 'DI0.2'
   TextField "Text field_20" at 244,258 size 22x53; Text 'DI0.3'
   TextField "Text field_21" at 272,258 size 22x53; Text 'DI0.4'
   TextField "Text field_22" at 300,258 size 22x53; Text 'DI0.5'
   TextField "Text field_23" at 328,258 size 22x53; Text 'DI0.6'
   TextField "Text field_24" at 356,258 size 22x53; Text 'DI0.7'
   TextField "Text field_25" at 404,258 size 22x53; Text 'DI1.0'
   TextField "Text field_26" at 432,258 size 22x53; Text 'DI1.1'
   TextField "Text field_27" at 460,258 size 22x53; Text 'DI1.2'
   TextField "Text field_28" at 488,258 size 22x53; Text 'DI1.3'
   TextField "Text field_29" at 516,258 size 22x53; Text 'DI1.4'
   TextField "Text field_30" at 544,258 size 22x53; Text 'DI1.5'
   TextField "Text field_31" at 572,258 size 22x53; Text 'DI1.6'
   TextField "Text field_32" at 600,258 size 22x53; Text 'DI1.7'
   TextField "Text field_33" at 648,258 size 22x53; Text 'DI2.0'
   TextField "Text field_34" at 676,258 size 22x53; Text 'DI2.1'
   TextField "Text field_35" at 704,258 size 22x53; Text 'DI2.2'
   TextField "Text field_36" at 732,258 size 22x53; Text 'DI2.3'
   TextField "Text field_37" at 760,258 size 22x53; Text 'DI2.4'
   TextField "Text field_38" at 788,258 size 22x53; Text 'DI2.5'
   TextField "Text field_39" at 816,258 size 22x53; Text 'DI2.6'
   TextField "Text field_40" at 844,258 size 22x53; Text 'DI2.7'
   TextField "Text field_41" at 892,258 size 22x53; Text 'DI3.0'
   TextField "Text field_42" at 920,258 size 22x53; Text 'DI3.1'
   TextField "Text field_43" at 948,258 size 22x53; Text 'DI3.2'
   TextField "Text field_44" at 976,258 size 22x53; Text 'DI3.3'
   TextField "Text field_45" at 1004,258 size 22x53; Text 'DI3.4'
   TextField "Text field_46" at 1032,258 size 22x53; Text 'DI3.5'
   TextField "Text field_47" at 1060,258 size 22x53; Text 'DI3.6'
   TextField "Text field_48" at 1088,258 size 22x53; Text 'DI3.7'
   TextField "Text field_49" at 158,572 size 22x58; Text 'DO0.0'
   TextField "Text field_50" at 186,572 size 22x58; Text 'DO0.1'
   TextField "Text field_51" at 214,572 size 22x58; Text 'DO0.2'
   TextField "Text field_52" at 242,572 size 22x58; Text 'DO0.3'
   TextField "Text field_53" at 270,572 size 22x58; Text 'DO0.4'
   TextField "Text field_54" at 298,572 size 22x58; Text 'DO0.5'
   TextField "Text field_55" at 326,572 size 22x58; Text 'DO0.6'
   TextField "Text field_56" at 354,572 size 22x58; Text 'DO0.7'
   TextField "Text field_57" at 402,572 size 22x58; Text 'DO1.0'
   TextField "Text field_58" at 430,572 size 22x58; Text 'DO1.1'
   TextField "Text field_59" at 458,572 size 22x58; Text 'DO1.2'
   TextField "Text field_60" at 486,572 size 22x58; Text 'DO1.3'
   TextField "Text field_61" at 514,572 size 22x58; Text 'DO1.4'
   TextField "Text field_62" at 542,572 size 22x58; Text 'DO1.5'
   TextField "Text field_63" at 570,572 size 22x58; Text 'DO1.6'
   TextField "Text field_64" at 598,572 size 22x58; Text 'DO1.7'
   TextField "Text field_65" at 646,572 size 22x58; Text 'DO2.0'
   TextField "Text field_66" at 674,572 size 22x58; Text 'DO2.1'
   TextField "Text field_67" at 702,572 size 22x58; Text 'DO2.2'
   TextField "Text field_68" at 730,572 size 22x58; Text 'DO2.3'
   TextField "Text field_69" at 758,572 size 22x58; Text 'DO2.4'
   TextField "Text field_70" at 786,572 size 22x58; Text 'DO2.5'
   TextField "Text field_71" at 814,572 size 22x58; Text 'DO2.6'
   TextField "Text field_72" at 842,572 size 22x58; Text 'DO2.7'
   TextField "Text field_73" at 890,572 size 22x58; Text 'DO3.0'
   TextField "Text field_74" at 918,572 size 22x58; Text 'DO3.1'
   TextField "Text field_75" at 946,572 size 22x58; Text 'DO3.2'
   TextField "Text field_76" at 974,572 size 22x58; Text 'DO3.3'
   TextField "Text field_77" at 1002,572 size 22x58; Text 'DO3.4'
   TextField "Text field_78" at 1030,572 size 22x58; Text 'DO3.5'
   TextField "Text field_79" at 1058,572 size 22x58; Text 'DO3.6'
   TextField "Text field_80" at 1086,572 size 22x58; Text 'DO3.7'

